REGION Network 68: CV60 PID TM_LAG
   RUNG wire#powerrail
      Contact( "Epics_to_PLC".CV60_PID_TM_LAG.cmdSet )
      { S7_GenerateENO := "TRUE" } Move(in := "Epics_to_PLC".CV60_PID_TM_LAG.cSetV, out1 => "PLC_to_Epics".CV60_PID_TM_LAG.sSetV)
      { S7_Templates := "SrcType := Real"; S7_GenerateENO := "TRUE" } Mul(in1 := "PLC_to_Epics".CV60_PID_TM_LAG.sSetV, in2 := 1000.0, out => #tmpR)
      { S7_Templates := "[SrcType := Real, DestType := DInt]"; S7_GenerateENO := "TRUE" } Round(in := #tmpR, out => "S4_Parameters".CV60_PID_TM_LAG)
      R_Coil( "Epics_to_PLC".CV60_PID_TM_LAG.cmdSet )
   END_RUNG
   // the same network as SCL:
   // ENO of a box is taken as its EN; it also drops when the box reports an error
   IF "Epics_to_PLC".CV60_PID_TM_LAG.cmdSet THEN
       "PLC_to_Epics".CV60_PID_TM_LAG.sSetV := "Epics_to_PLC".CV60_PID_TM_LAG.cSetV;
       #tmpR := "PLC_to_Epics".CV60_PID_TM_LAG.sSetV * 1000.0;
       "S4_Parameters".CV60_PID_TM_LAG := ROUND(#tmpR);
       "Epics_to_PLC".CV60_PID_TM_LAG.cmdSet := FALSE;
   END_IF;
END_REGION
END_FUNCTION

FUNCTION "Data_from_IOC" : Void   // FC34, LAD
TITLE = Get data from the IOC andcheck if the connection is alive
{ S7_Optimized_Access := 'FALSE' }
VERSION : 0.1
BEGIN

REGION Network 1: Check the Data from the IOC
END_REGION
END_FUNCTION

FUNCTION "grafcet" : Void   // FC99, LAD
{ S7_Optimized_Access := 'FALSE' }
VERSION : 0.1
   VAR_TEMP   // added for the SCL form of the ladder/FBD networks
      _w1 : Bool;
      _w2 : Bool;
      _w3 : Bool;
      _w4 : Bool;
      _w5 : Bool;
      _w6 : Bool;
      _w7 : Bool;
      _w8 : Bool;
   END_VAR
BEGIN

REGION Network 1: Set initial step number for the state S4
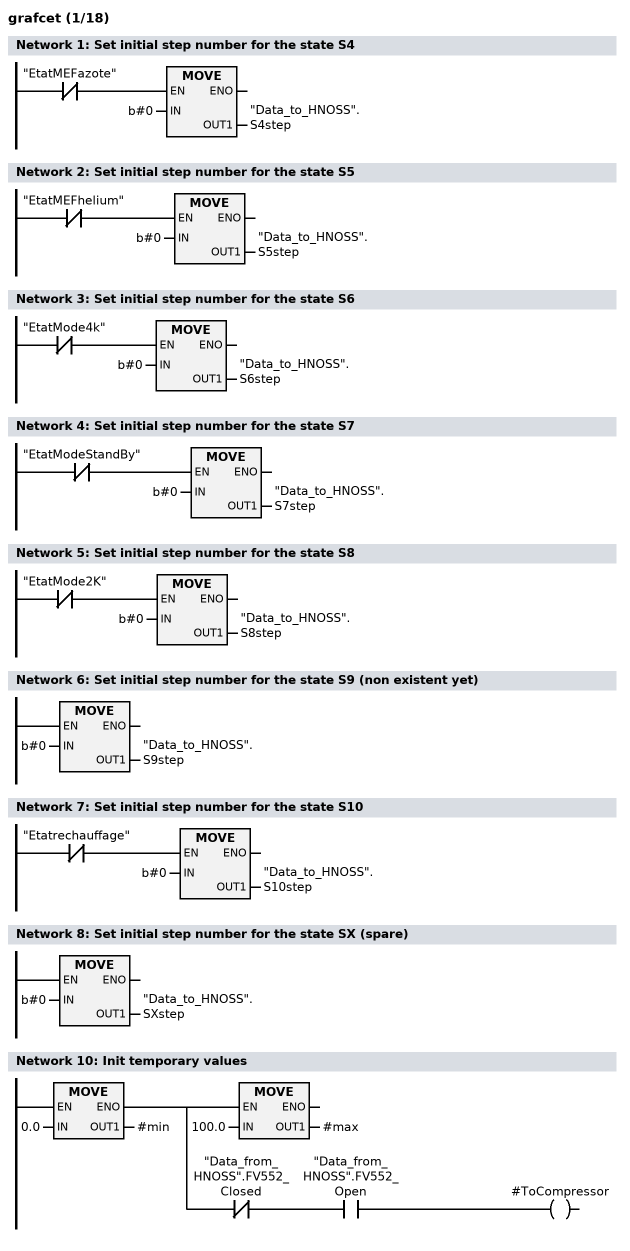
   RUNG wire#powerrail
      I_Contact( "EtatMEFazote" )
      { S7_GenerateENO := "TRUE" } Move(in := b#0, out1 => "Data_to_HNOSS".S4step)
   END_RUNG
   // the same network as SCL:
   IF NOT "EtatMEFazote" THEN "Data_to_HNOSS".S4step := b#0; END_IF;
END_REGION

REGION Network 2: Set initial step number for the state S5
   RUNG wire#powerrail
      I_Contact( "EtatMEFhelium" )
      { S7_GenerateENO := "TRUE" } Move(in := b#0, out1 => "Data_to_HNOSS".S5step)
   END_RUNG
   // the same network as SCL:
   IF NOT "EtatMEFhelium" THEN "Data_to_HNOSS".S5step := b#0; END_IF;
END_REGION

REGION Network 3: Set initial step number for the state S6
   RUNG wire#powerrail
      I_Contact( "EtatMode4k" )
      { S7_GenerateENO := "TRUE" } Move(in := b#0, out1 => "Data_to_HNOSS".S6step)
   END_RUNG
   // the same network as SCL:
   IF NOT "EtatMode4k" THEN "Data_to_HNOSS".S6step := b#0; END_IF;
END_REGION

REGION Network 4: Set initial step number for the state S7
   RUNG wire#powerrail
      I_Contact( "EtatModeStandBy" )
      { S7_GenerateENO := "TRUE" } Move(in := b#0, out1 => "Data_to_HNOSS".S7step)
   END_RUNG
   // the same network as SCL:
   IF NOT "EtatModeStandBy" THEN "Data_to_HNOSS".S7step := b#0; END_IF;
END_REGION

REGION Network 5: Set initial step number for the state S8
   RUNG wire#powerrail
      I_Contact( "EtatMode2K" )
      { S7_GenerateENO := "TRUE" } Move(in := b#0, out1 => "Data_to_HNOSS".S8step)
   END_RUNG
   // the same network as SCL:
   IF NOT "EtatMode2K" THEN "Data_to_HNOSS".S8step := b#0; END_IF;
END_REGION

REGION Network 6: Set initial step number for the state S9 (non existent yet)
   RUNG wire#powerrail
      { S7_GenerateENO := "TRUE" } Move(in := b#0, out1 => "Data_to_HNOSS".S9step)
   END_RUNG
   // the same network as SCL:
   "Data_to_HNOSS".S9step := b#0;
END_REGION

REGION Network 7: Set initial step number for the state S10
   RUNG wire#powerrail
      I_Contact( "Etatrechauffage" )
      { S7_GenerateENO := "TRUE" } Move(in := b#0, out1 => "Data_to_HNOSS".S10step)
   END_RUNG
   // the same network as SCL:
   IF NOT "Etatrechauffage" THEN "Data_to_HNOSS".S10step := b#0; END_IF;
END_REGION

REGION Network 8: Set initial step number for the state SX (spare)
   RUNG wire#powerrail
      { S7_GenerateENO := "TRUE" } Move(in := b#0, out1 => "Data_to_HNOSS".SXstep)
   END_RUNG
   // the same network as SCL:
   "Data_to_HNOSS".SXstep := b#0;
END_REGION

REGION Network 9 (STL): Change to int for "compare" instruction

         L     "Data_to_HNOSS".S4step;
         T     #S4step;
         L     "Data_to_HNOSS".S5step;
         T     #S5step;
         L     "Data_to_HNOSS".S6step;
         T     #S6step;
         L     "Data_to_HNOSS".S7step;
         T     #S7step;
         L     "Data_to_HNOSS".S8step;
         T     #S8step;
         L     "Data_to_HNOSS".S9step;
         T     #S9step;
         L     "Data_to_HNOSS".S10step;
         T     #S10step;
         L     "Data_to_HNOSS".SXstep;
         T     #Sxstep;
END_REGION

REGION Network 10: Init temporary values
   RUNG wire#powerrail
      { S7_GenerateENO := "TRUE" } Move(in := 0.0, out1 => #min)
      wire#w1
      { S7_GenerateENO := "TRUE" } Move(in := 100.0, out1 => #max)
   END_RUNG
   RUNG wire#w1
      I_Contact( "Data_from_HNOSS".FV552_Closed )
      Contact( "Data_from_HNOSS".FV552_Open )
      Coil( #ToCompressor )
   END_RUNG
   // the same network as SCL:
   // ENO of a box is taken as its EN; it also drops when the box reports an error
   #min := 0.0;
   #max := 100.0;
   #ToCompressor := NOT "Data_from_HNOSS".FV552_Closed AND "Data_from_HNOSS".FV552_Open;
END_REGION

REGION Network 11: config vannes init mode
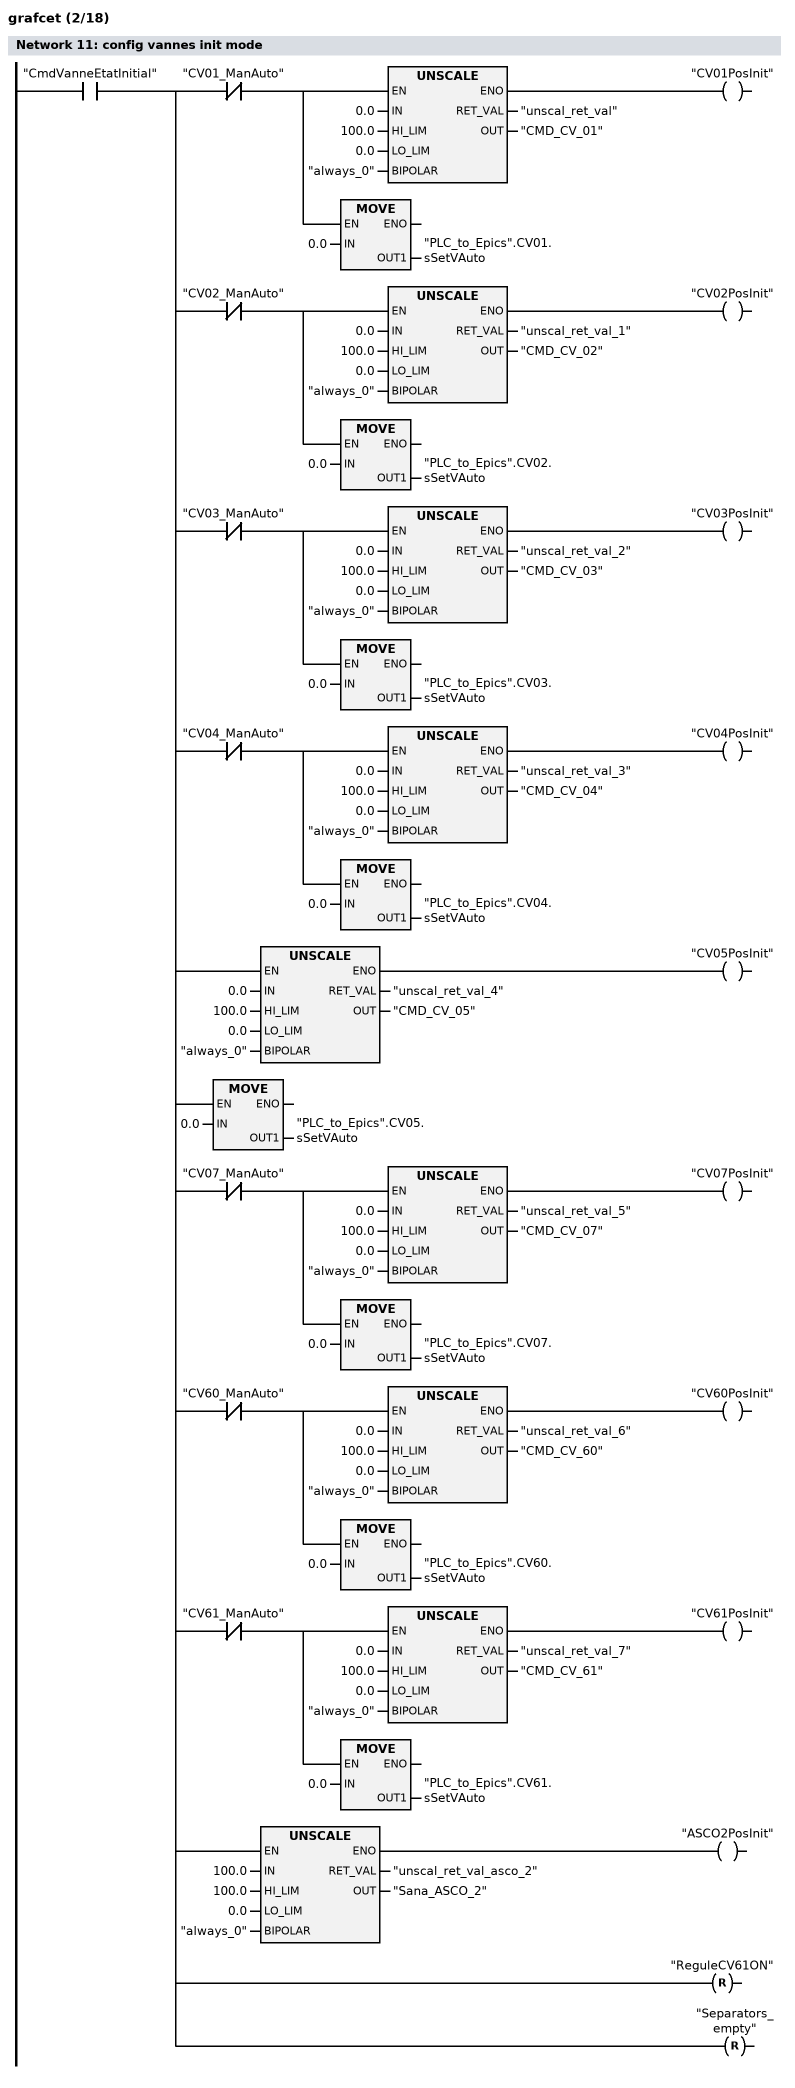
   // ENO of a box is taken as its EN; it also drops when the box reports an error
   #_w1 := "CmdVanneEtatInitial" AND NOT "CV01_ManAuto";
   #_w2 := "CmdVanneEtatInitial";
   IF #_w1 THEN
       "unscal_ret_val" := UNSCALE(IN := 0.0,
                               HI_LIM := 100.0,
                               LO_LIM := 0.0,
                               BIPOLAR := "always_0",
                               OUT => "CMD_CV_01");
   END_IF;
   "CV01PosInit" := #_w1;
   IF #_w1 THEN "PLC_to_Epics".CV01.sSetVAuto := 0.0; END_IF;
   #_w3 := #_w2 AND NOT "CV02_ManAuto";
   IF #_w3 THEN
       "unscal_ret_val_1" := UNSCALE(IN := 0.0,
                               HI_LIM := 100.0,
                               LO_LIM := 0.0,
                               BIPOLAR := "always_0",
                               OUT => "CMD_CV_02");
   END_IF;
   "CV02PosInit" := #_w3;
   IF #_w3 THEN "PLC_to_Epics".CV02.sSetVAuto := 0.0; END_IF;
   #_w4 := #_w2 AND NOT "CV03_ManAuto";
   IF #_w4 THEN
       "unscal_ret_val_2" := UNSCALE(IN := 0.0,
                               HI_LIM := 100.0,
                               LO_LIM := 0.0,
                               BIPOLAR := "always_0",
                               OUT => "CMD_CV_03");
   END_IF;
   "CV03PosInit" := #_w4;
   IF #_w4 THEN "PLC_to_Epics".CV03.sSetVAuto := 0.0; END_IF;
   #_w5 := #_w2 AND NOT "CV04_ManAuto";
   IF #_w5 THEN
       "unscal_ret_val_3" := UNSCALE(IN := 0.0,
                               HI_LIM := 100.0,
                               LO_LIM := 0.0,
                               BIPOLAR := "always_0",
                               OUT => "CMD_CV_04");
   END_IF;
   "CV04PosInit" := #_w5;
   IF #_w5 THEN "PLC_to_Epics".CV04.sSetVAuto := 0.0; END_IF;
   IF #_w2 THEN
       "unscal_ret_val_4" := UNSCALE(IN := 0.0,
                               HI_LIM := 100.0,
                               LO_LIM := 0.0,
                               BIPOLAR := "always_0",
                               OUT => "CMD_CV_05");
   END_IF;
   "CV05PosInit" := #_w2;
   IF #_w2 THEN "PLC_to_Epics".CV05.sSetVAuto := 0.0; END_IF;
   #_w6 := #_w2 AND NOT "CV07_ManAuto";
   IF #_w6 THEN
       "unscal_ret_val_5" := UNSCALE(IN := 0.0,
                               HI_LIM := 100.0,
                               LO_LIM := 0.0,
                               BIPOLAR := "always_0",
                               OUT => "CMD_CV_07");
   END_IF;
   "CV07PosInit" := #_w6;
   IF #_w6 THEN "PLC_to_Epics".CV07.sSetVAuto := 0.0; END_IF;
   #_w7 := #_w2 AND NOT "CV60_ManAuto";
   IF #_w7 THEN
       "unscal_ret_val_6" := UNSCALE(IN := 0.0,
                               HI_LIM := 100.0,
                               LO_LIM := 0.0,
                               BIPOLAR := "always_0",
                               OUT => "CMD_CV_60");
   END_IF;
   "CV60PosInit" := #_w7;
   IF #_w7 THEN "PLC_to_Epics".CV60.sSetVAuto := 0.0; END_IF;
   #_w8 := #_w2 AND NOT "CV61_ManAuto";
   IF #_w8 THEN
       "unscal_ret_val_7" := UNSCALE(IN := 0.0,
                               HI_LIM := 100.0,
                               LO_LIM := 0.0,
                               BIPOLAR := "always_0",
                               OUT => "CMD_CV_61");
   END_IF;
   "CV61PosInit" := #_w8;
   IF #_w8 THEN "PLC_to_Epics".CV61.sSetVAuto := 0.0; END_IF;
   IF #_w2 THEN
       "unscal_ret_val_asco_2" := UNSCALE(IN := 100.0,
                               HI_LIM := 100.0,
                               LO_LIM := 0.0,
                               BIPOLAR := "always_0",
                               OUT => "Sana_ASCO_2");
   END_IF;
   "ASCO2PosInit" := #_w2;
   IF #_w2 THEN
       "ReguleCV61ON" := FALSE;
       "Separators_empty" := FALSE;
   END_IF;
END_REGION

REGION Network 12: Vanne En Position Initial
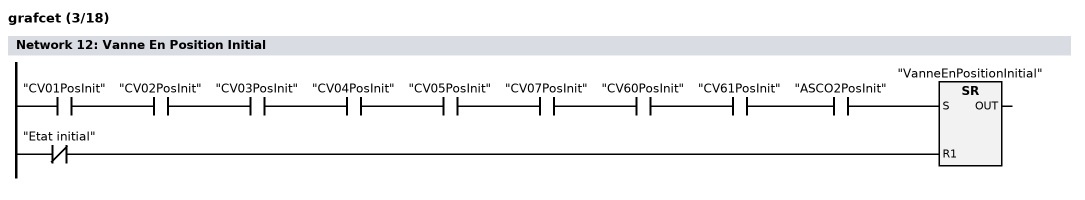
   RUNG wire#powerrail
      Contact( "CV01PosInit" )
      Contact( "CV02PosInit" )
      Contact( "CV03PosInit" )
      Contact( "CV04PosInit" )
      Contact( "CV05PosInit" )
      Contact( "CV07PosInit" )
      Contact( "CV60PosInit" )
      Contact( "CV61PosInit" )
      Contact( "ASCO2PosInit" )
      S_SR(operand := "VanneEnPositionInitial", r1 := wire#w1)
   END_RUNG
   RUNG wire#powerrail
      I_Contact( "Etat initial" )
   END_RUNG wire#w1
   // the same network as SCL:
   IF "CV01PosInit" AND "CV02PosInit" AND "CV03PosInit" AND "CV04PosInit" AND "CV05PosInit" AND "CV07PosInit" AND "CV60PosInit" AND "CV61PosInit" AND "ASCO2PosInit" THEN
       "VanneEnPositionInitial" := TRUE;   // SR flip-flop
   END_IF;
   IF NOT "Etat initial" THEN "VanneEnPositionInitial" := FALSE; END_IF;
END_REGION

REGION Network 13: config vanne etat conditionnement
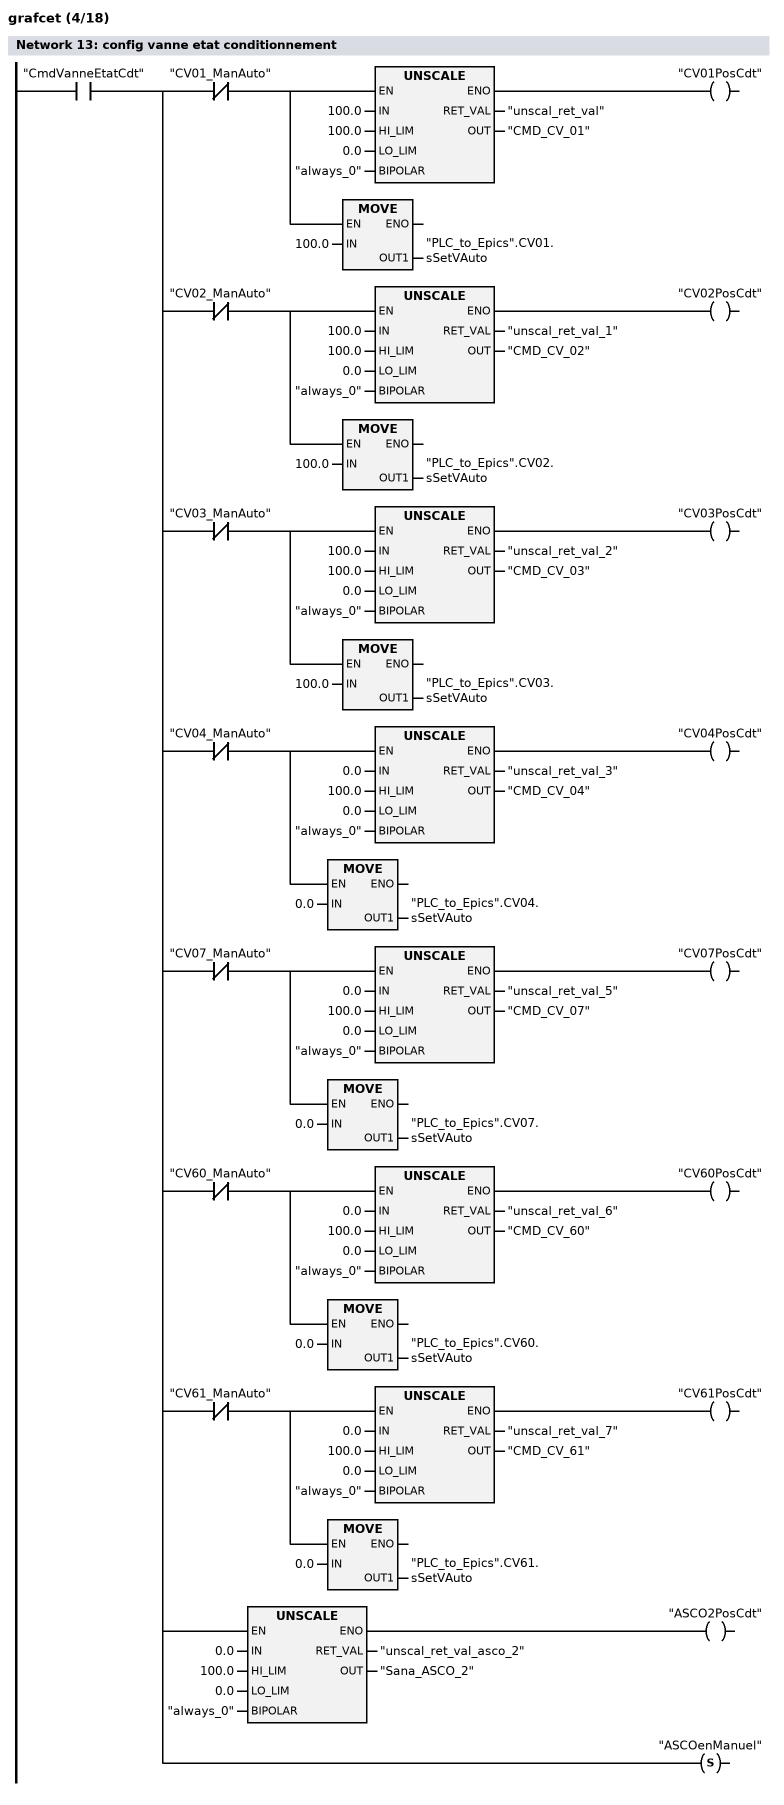
   // ENO of a box is taken as its EN; it also drops when the box reports an error
   #_w1 := "CmdVanneEtatCdt" AND NOT "CV01_ManAuto";
   #_w2 := "CmdVanneEtatCdt";
   IF #_w1 THEN
       "unscal_ret_val" := UNSCALE(IN := 100.0,
                               HI_LIM := 100.0,
                               LO_LIM := 0.0,
                               BIPOLAR := "always_0",
                               OUT => "CMD_CV_01");
   END_IF;
   "CV01PosCdt" := #_w1;
   IF #_w1 THEN "PLC_to_Epics".CV01.sSetVAuto := 100.0; END_IF;
   #_w3 := #_w2 AND NOT "CV02_ManAuto";
   IF #_w3 THEN
       "unscal_ret_val_1" := UNSCALE(IN := 100.0,
                               HI_LIM := 100.0,
                               LO_LIM := 0.0,
                               BIPOLAR := "always_0",
                               OUT => "CMD_CV_02");
   END_IF;
   "CV02PosCdt" := #_w3;
   IF #_w3 THEN "PLC_to_Epics".CV02.sSetVAuto := 100.0; END_IF;
   #_w4 := #_w2 AND NOT "CV03_ManAuto";
   IF #_w4 THEN
       "unscal_ret_val_2" := UNSCALE(IN := 100.0,
                               HI_LIM := 100.0,
                               LO_LIM := 0.0,
                               BIPOLAR := "always_0",
                               OUT => "CMD_CV_03");
   END_IF;
   "CV03PosCdt" := #_w4;
   IF #_w4 THEN "PLC_to_Epics".CV03.sSetVAuto := 100.0; END_IF;
   #_w5 := #_w2 AND NOT "CV04_ManAuto";
   IF #_w5 THEN
       "unscal_ret_val_3" := UNSCALE(IN := 0.0,
                               HI_LIM := 100.0,
                               LO_LIM := 0.0,
                               BIPOLAR := "always_0",
                               OUT => "CMD_CV_04");
   END_IF;
   "CV04PosCdt" := #_w5;
   IF #_w5 THEN "PLC_to_Epics".CV04.sSetVAuto := 0.0; END_IF;
   #_w6 := #_w2 AND NOT "CV07_ManAuto";
   IF #_w6 THEN
       "unscal_ret_val_5" := UNSCALE(IN := 0.0,
                               HI_LIM := 100.0,
                               LO_LIM := 0.0,
                               BIPOLAR := "always_0",
                               OUT => "CMD_CV_07");
   END_IF;
   "CV07PosCdt" := #_w6;
   IF #_w6 THEN "PLC_to_Epics".CV07.sSetVAuto := 0.0; END_IF;
   #_w7 := #_w2 AND NOT "CV60_ManAuto";
   IF #_w7 THEN
       "unscal_ret_val_6" := UNSCALE(IN := 0.0,
                               HI_LIM := 100.0,
                               LO_LIM := 0.0,
                               BIPOLAR := "always_0",
                               OUT => "CMD_CV_60");
   END_IF;
   "CV60PosCdt" := #_w7;
   IF #_w7 THEN "PLC_to_Epics".CV60.sSetVAuto := 0.0; END_IF;
   #_w8 := #_w2 AND NOT "CV61_ManAuto";
   IF #_w8 THEN
       "unscal_ret_val_7" := UNSCALE(IN := 0.0,
                               HI_LIM := 100.0,
                               LO_LIM := 0.0,
                               BIPOLAR := "always_0",
                               OUT => "CMD_CV_61");
   END_IF;
   "CV61PosCdt" := #_w8;
   IF #_w8 THEN "PLC_to_Epics".CV61.sSetVAuto := 0.0; END_IF;
   IF #_w2 THEN
       "unscal_ret_val_asco_2" := UNSCALE(IN := 0.0,
                               HI_LIM := 100.0,
                               LO_LIM := 0.0,
                               BIPOLAR := "always_0",
                               OUT => "Sana_ASCO_2");
   END_IF;
   "ASCO2PosCdt" := #_w2;
   IF #_w2 THEN "ASCOenManuel" := TRUE; END_IF;
END_REGION

REGION Network 14: Vanne En Position Cdt
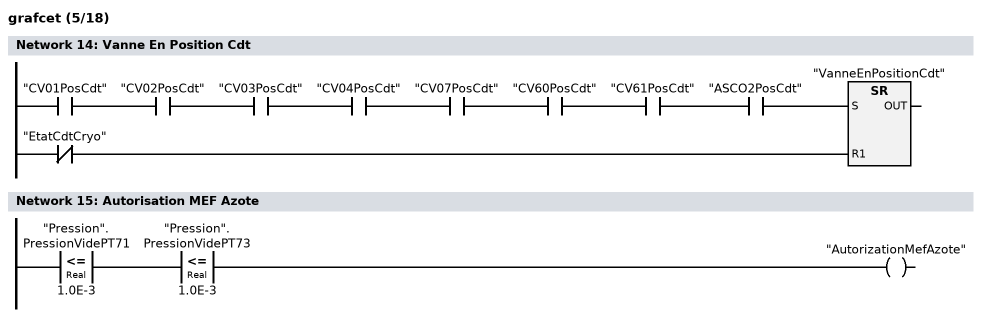
   RUNG wire#powerrail
      Contact( "CV01PosCdt" )
      Contact( "CV02PosCdt" )
      Contact( "CV03PosCdt" )
      Contact( "CV04PosCdt" )
      Contact( "CV07PosCdt" )
      Contact( "CV60PosCdt" )
      Contact( "CV61PosCdt" )
      Contact( "ASCO2PosCdt" )
      S_SR(operand := "VanneEnPositionCdt", r1 := wire#w1)
   END_RUNG
   RUNG wire#powerrail
      I_Contact( "EtatCdtCryo" )
   END_RUNG wire#w1
   // the same network as SCL:
   IF "CV01PosCdt" AND "CV02PosCdt" AND "CV03PosCdt" AND "CV04PosCdt" AND "CV07PosCdt" AND "CV60PosCdt" AND "CV61PosCdt" AND "ASCO2PosCdt" THEN
       "VanneEnPositionCdt" := TRUE;   // SR flip-flop
   END_IF;
   IF NOT "EtatCdtCryo" THEN "VanneEnPositionCdt" := FALSE; END_IF;
END_REGION

REGION Network 15: Autorisation MEF Azote
   RUNG wire#powerrail
      { S7_Templates := "SrcType := Real" } LE_Contact(in1 := "Pression".PressionVidePT71, in2 := 1.0E-3)
      { S7_Templates := "SrcType := Real" } LE_Contact(in1 := "Pression".PressionVidePT73, in2 := 1.0E-3)
      Coil( "AutorizationMefAzote" )
   END_RUNG
   // the same network as SCL:
   "AutorizationMefAzote" := ("Pression".PressionVidePT71 <= 1.0E-3) AND ("Pression".PressionVidePT73 <= 1.0E-3);
END_REGION

REGION Network 16: config vannes init mode & regule cv61 on
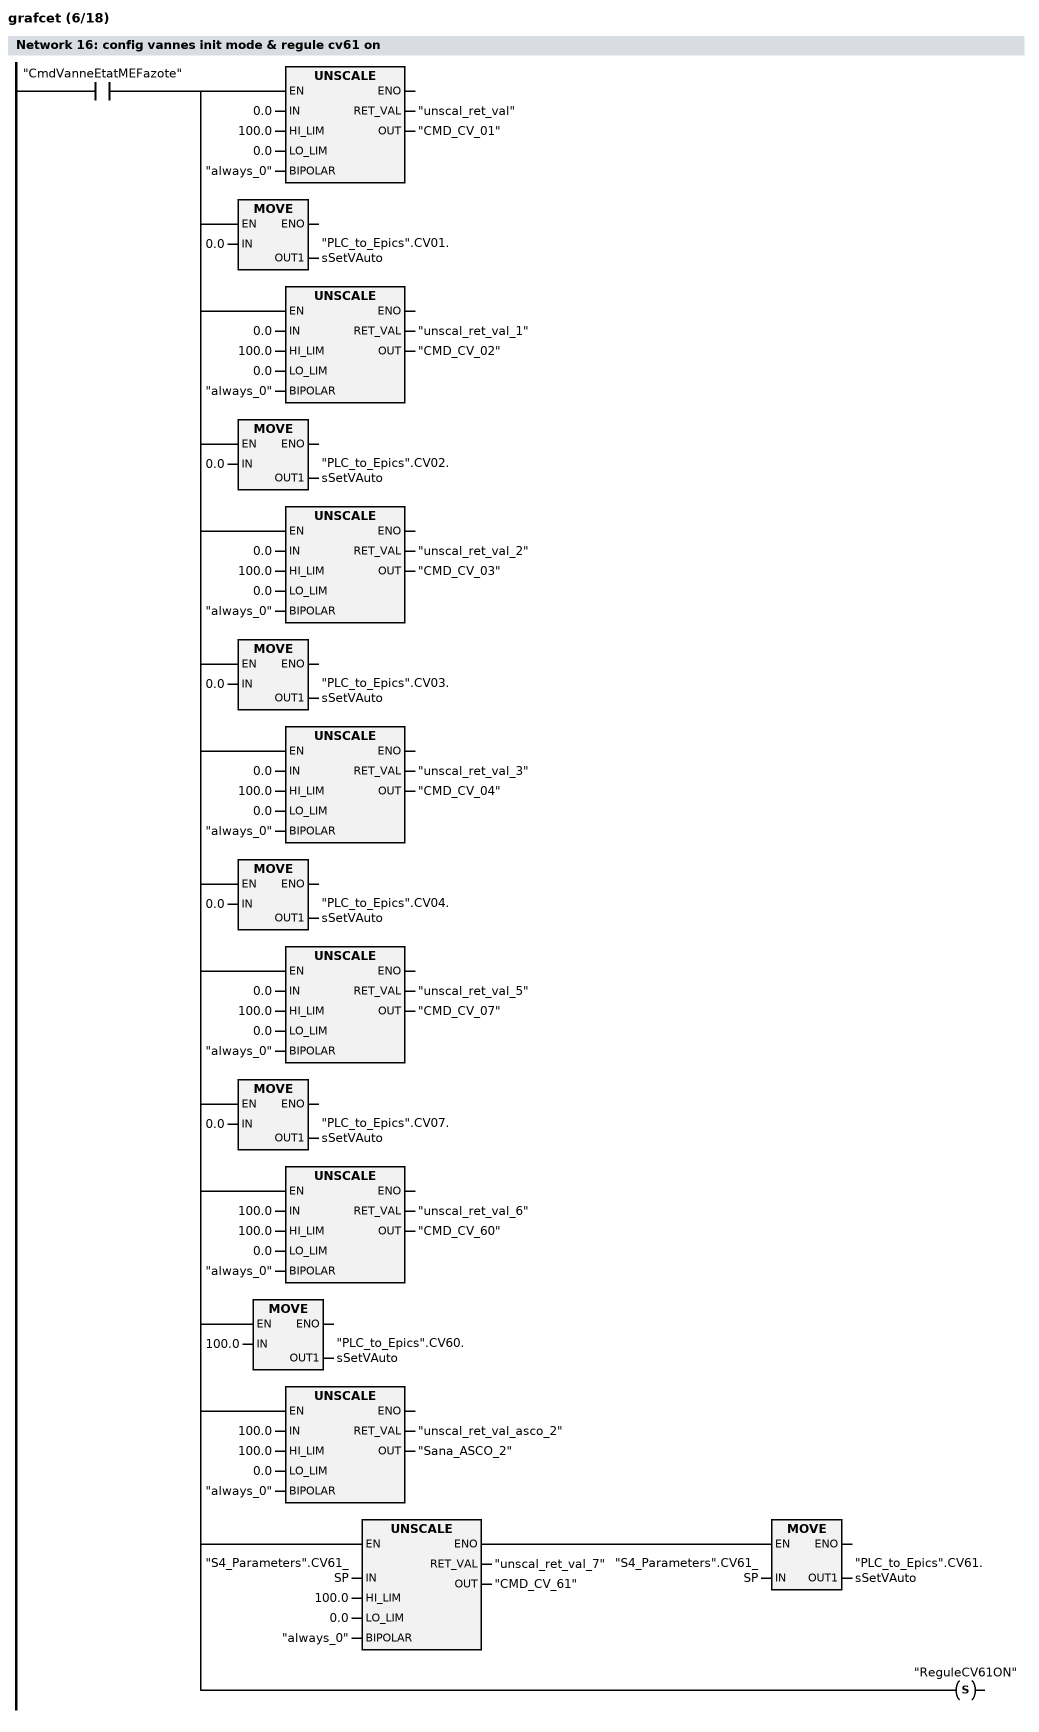
   // ENO of a box is taken as its EN; it also drops when the box reports an error
   #_w1 := "CmdVanneEtatMEFazote";
   IF #_w1 THEN
       "unscal_ret_val" := UNSCALE(IN := 0.0,
                               HI_LIM := 100.0,
                               LO_LIM := 0.0,
                               BIPOLAR := "always_0",
                               OUT => "CMD_CV_01");
       "PLC_to_Epics".CV01.sSetVAuto := 0.0;
       "unscal_ret_val_1" := UNSCALE(IN := 0.0,
                               HI_LIM := 100.0,
                               LO_LIM := 0.0,
                               BIPOLAR := "always_0",
                               OUT => "CMD_CV_02");
       "PLC_to_Epics".CV02.sSetVAuto := 0.0;
       "unscal_ret_val_2" := UNSCALE(IN := 0.0,
                               HI_LIM := 100.0,
                               LO_LIM := 0.0,
                               BIPOLAR := "always_0",
                               OUT => "CMD_CV_03");
       "PLC_to_Epics".CV03.sSetVAuto := 0.0;
       "unscal_ret_val_3" := UNSCALE(IN := 0.0,
                               HI_LIM := 100.0,
                               LO_LIM := 0.0,
                               BIPOLAR := "always_0",
                               OUT => "CMD_CV_04");
       "PLC_to_Epics".CV04.sSetVAuto := 0.0;
       "unscal_ret_val_5" := UNSCALE(IN := 0.0,
                               HI_LIM := 100.0,
                               LO_LIM := 0.0,
                               BIPOLAR := "always_0",
                               OUT => "CMD_CV_07");
       "PLC_to_Epics".CV07.sSetVAuto := 0.0;
       "unscal_ret_val_6" := UNSCALE(IN := 100.0,
                               HI_LIM := 100.0,
                               LO_LIM := 0.0,
                               BIPOLAR := "always_0",
                               OUT => "CMD_CV_60");
       "PLC_to_Epics".CV60.sSetVAuto := 100.0;
       "unscal_ret_val_asco_2" := UNSCALE(IN := 100.0,
                               HI_LIM := 100.0,
                               LO_LIM := 0.0,
                               BIPOLAR := "always_0",
                               OUT => "Sana_ASCO_2");
       "unscal_ret_val_7" := UNSCALE(IN := "S4_Parameters".CV61_SP,
                               HI_LIM := 100.0,
                               LO_LIM := 0.0,
                               BIPOLAR := "always_0",
                               OUT => "CMD_CV_61");
       "PLC_to_Epics".CV61.sSetVAuto := "S4_Parameters".CV61_SP;
       "ReguleCV61ON" := TRUE;
   END_IF;
END_REGION

REGION Network 17: Régule CV61 seuil (desactive)
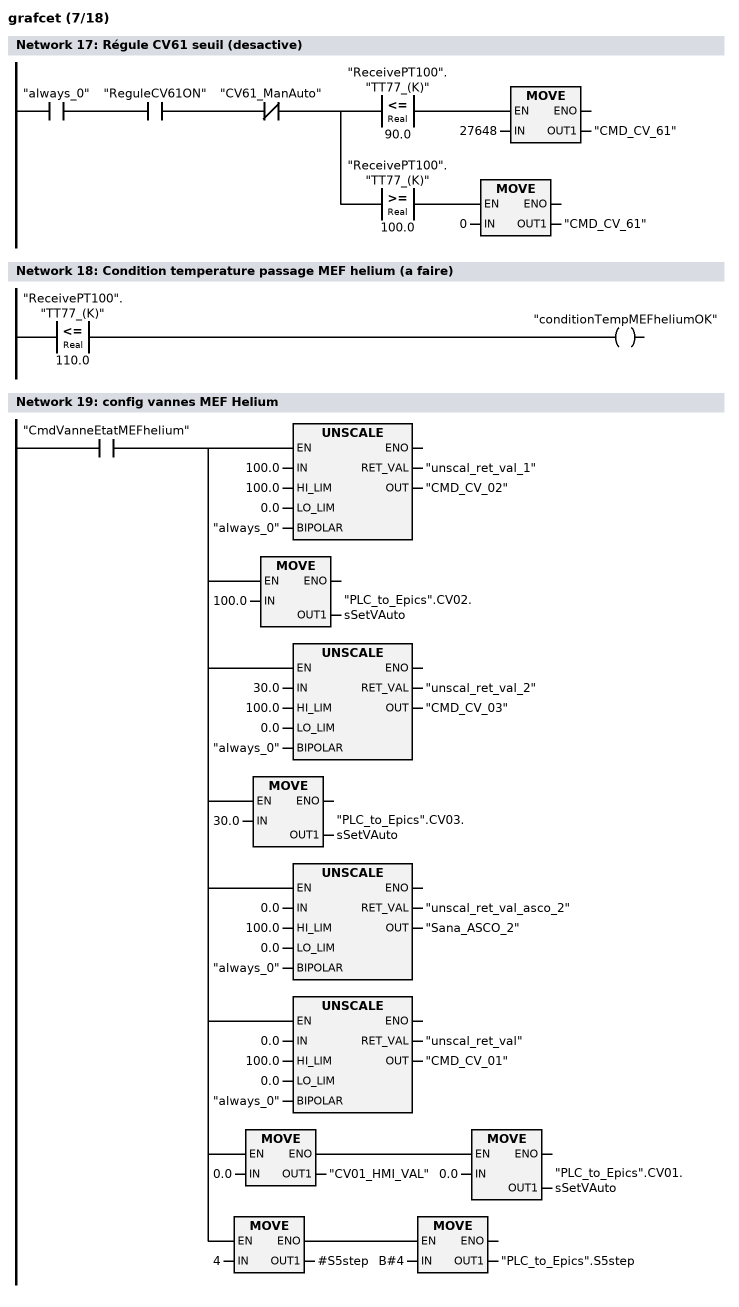
   RUNG wire#powerrail
      Contact( "always_0" )
      Contact( "ReguleCV61ON" )
      I_Contact( "CV61_ManAuto" )
      wire#w1
      { S7_Templates := "SrcType := Real" } LE_Contact(in1 := "ReceivePT100"."TT77_(K)", in2 := 90.0)
      { S7_GenerateENO := "TRUE" } Move(in := 27648, out1 => "CMD_CV_61")
   END_RUNG
   RUNG wire#w1
      { S7_Templates := "SrcType := Real" } GE_Contact(in1 := "ReceivePT100"."TT77_(K)", in2 := 100.0)
      { S7_GenerateENO := "TRUE" } Move(in := 0, out1 => "CMD_CV_61")
   END_RUNG
   // the same network as SCL:
   #_w1 := "always_0" AND "ReguleCV61ON" AND NOT "CV61_ManAuto";
   IF #_w1 AND ("ReceivePT100"."TT77_(K)" <= 90.0) THEN "CMD_CV_61" := 27648; END_IF;
   IF #_w1 AND ("ReceivePT100"."TT77_(K)" >= 100.0) THEN "CMD_CV_61" := 0; END_IF;
END_REGION

REGION Network 18: Condition temperature passage MEF helium (a faire)
   RUNG wire#powerrail
      { S7_Templates := "SrcType := Real" } LE_Contact(in1 := "ReceivePT100"."TT77_(K)", in2 := 110.0)
      Coil( "conditionTempMEFheliumOK" )
   END_RUNG
   // the same network as SCL:
   "conditionTempMEFheliumOK" := "ReceivePT100"."TT77_(K)" <= 110.0;
END_REGION

REGION Network 19: config vannes MEF Helium
   // ENO of a box is taken as its EN; it also drops when the box reports an error
   #_w1 := "CmdVanneEtatMEFhelium";
   IF #_w1 THEN
       "unscal_ret_val_1" := UNSCALE(IN := 100.0,
                               HI_LIM := 100.0,
                               LO_LIM := 0.0,
                               BIPOLAR := "always_0",
                               OUT => "CMD_CV_02");
       "PLC_to_Epics".CV02.sSetVAuto := 100.0;
       "unscal_ret_val_2" := UNSCALE(IN := 30.0,
                               HI_LIM := 100.0,
                               LO_LIM := 0.0,
                               BIPOLAR := "always_0",
                               OUT => "CMD_CV_03");
       "PLC_to_Epics".CV03.sSetVAuto := 30.0;
       "unscal_ret_val_asco_2" := UNSCALE(IN := 0.0,
                               HI_LIM := 100.0,
                               LO_LIM := 0.0,
                               BIPOLAR := "always_0",
                               OUT => "Sana_ASCO_2");
       "unscal_ret_val" := UNSCALE(IN := 0.0,
                               HI_LIM := 100.0,
                               LO_LIM := 0.0,
                               BIPOLAR := "always_0",
                               OUT => "CMD_CV_01");
       "CV01_HMI_VAL" := 0.0;
       "PLC_to_Epics".CV01.sSetVAuto := 0.0;
       #S5step := 4;
       "PLC_to_Epics".S5step := B#4;
   END_IF;
END_REGION

REGION Network 20: LHe cooling down - Set step 6 (maybe setting CV03 is not needed here (done in the next network)!!!!!